       //Move FIRE HMW
       //H1
       "M256_Manag_IDB".M256F_IDB[0].tHMW.dHeadFireONReaction_ms := "DB_M256F_Scada".tHMW.dHeadFireONReaction_ms_H1;
       "M256_Manag_IDB".M256F_IDB[0].tHMW.dHeadFireOFFReaction_ms := "DB_M256F_Scada".tHMW.dHeadFireOFFReaction_ms_H1;
       "M256_Manag_IDB".M256F_IDB[0].tHMW.dHeadOilONDelay_ms := "DB_M256F_Scada".tHMW.dHeadOilONDelay_ms_H1;
       "M256_Manag_IDB".M256F_IDB[0].tHMW.dHeadOilOFFDelay_ms := "DB_M256F_Scada".tHMW.dHeadOilOFFDelay_ms_H1;
       "M256_Manag_IDB".M256F_IDB[0].tHMW.dHeadFireONDelay_cmm := "DB_M256F_Scada".tHMW.dHeadFireONDelay_cmm_H1;
       "M256_Manag_IDB".M256F_IDB[0].tHMW.dHeadFireOFFDelay_cmm := "DB_M256F_Scada".tHMW.dHeadFireOFFDelay_cmm_H1;
       "M256_Manag_IDB".M256F_IDB[0].tHMW.dHeadPressure_mN := "DB_M256F_Scada".tHMW.dHeadPressure_mN_H1;
       "M256_Manag_IDB".M256F_IDB[0].tHMW.xResetUsageCounter := "DB_M256F_Scada".tHMW.xResetUsageCounter_H1;
       "M256_Manag_IDB".M256F_IDB[0].tHMW.tManCmd.xMan_FireON := "DB_M256F_Scada".tHMW.tManCmd.xMan_FireON_H1;
       "M256_Manag_IDB".M256F_IDB[0].tHMW.tManCmd.xMan_FireOFF := "DB_M256F_Scada".tHMW.tManCmd.xMan_FireOFF_H1;
       "M256_Manag_IDB".M256F_IDB[0].tHMW.tManCmd.xMan_OilON := "DB_M256F_Scada".tHMW.tManCmd.xMan_OilON_H1;
       //H2
       "M256_Manag_IDB".M256F_IDB[1].tHMW.dHeadFireONReaction_ms := "DB_M256F_Scada".tHMW.dHeadFireONReaction_ms_H2;
       "M256_Manag_IDB".M256F_IDB[1].tHMW.dHeadFireOFFReaction_ms := "DB_M256F_Scada".tHMW.dHeadFireOFFReaction_ms_H2;
       "M256_Manag_IDB".M256F_IDB[1].tHMW.dHeadOilONDelay_ms := "DB_M256F_Scada".tHMW.dHeadOilONDelay_ms_H2;
       "M256_Manag_IDB".M256F_IDB[1].tHMW.dHeadOilOFFDelay_ms := "DB_M256F_Scada".tHMW.dHeadOilOFFDelay_ms_H2;
       "M256_Manag_IDB".M256F_IDB[1].tHMW.dHeadFireONDelay_cmm := "DB_M256F_Scada".tHMW.dHeadFireONDelay_cmm_H2;
       "M256_Manag_IDB".M256F_IDB[1].tHMW.dHeadFireOFFDelay_cmm := "DB_M256F_Scada".tHMW.dHeadFireOFFDelay_cmm_H2;
       "M256_Manag_IDB".M256F_IDB[1].tHMW.dHeadPressure_mN := "DB_M256F_Scada".tHMW.dHeadPressure_mN_H2;
       "M256_Manag_IDB".M256F_IDB[1].tHMW.xResetUsageCounter := "DB_M256F_Scada".tHMW.xResetUsageCounter_H2;
       "M256_Manag_IDB".M256F_IDB[1].tHMW.tManCmd.xMan_FireON := "DB_M256F_Scada".tHMW.tManCmd.xMan_FireON_H2;
       "M256_Manag_IDB".M256F_IDB[1].tHMW.tManCmd.xMan_FireOFF := "DB_M256F_Scada".tHMW.tManCmd.xMan_FireOFF_H2;
       "M256_Manag_IDB".M256F_IDB[1].tHMW.tManCmd.xMan_OilON := "DB_M256F_Scada".tHMW.tManCmd.xMan_OilON_H2;
       //H3
       "M256_Manag_IDB".M256F_IDB[2].tHMW.dHeadFireONReaction_ms := "DB_M256F_Scada".tHMW.dHeadFireONReaction_ms_H3;
       "M256_Manag_IDB".M256F_IDB[2].tHMW.dHeadFireOFFReaction_ms := "DB_M256F_Scada".tHMW.dHeadFireOFFReaction_ms_H3;
       "M256_Manag_IDB".M256F_IDB[2].tHMW.dHeadOilONDelay_ms := "DB_M256F_Scada".tHMW.dHeadOilONDelay_ms_H3;
       "M256_Manag_IDB".M256F_IDB[2].tHMW.dHeadOilOFFDelay_ms := "DB_M256F_Scada".tHMW.dHeadOilOFFDelay_ms_H3;
       "M256_Manag_IDB".M256F_IDB[2].tHMW.dHeadFireONDelay_cmm := "DB_M256F_Scada".tHMW.dHeadFireONDelay_cmm_H3;
       "M256_Manag_IDB".M256F_IDB[2].tHMW.dHeadFireOFFDelay_cmm := "DB_M256F_Scada".tHMW.dHeadFireOFFDelay_cmm_H3;
       "M256_Manag_IDB".M256F_IDB[2].tHMW.dHeadPressure_mN := "DB_M256F_Scada".tHMW.dHeadPressure_mN_H3;
       "M256_Manag_IDB".M256F_IDB[2].tHMW.xResetUsageCounter := "DB_M256F_Scada".tHMW.xResetUsageCounter_H3;
       "M256_Manag_IDB".M256F_IDB[2].tHMW.tManCmd.xMan_FireON := "DB_M256F_Scada".tHMW.tManCmd.xMan_FireON_H3;
       "M256_Manag_IDB".M256F_IDB[2].tHMW.tManCmd.xMan_FireOFF := "DB_M256F_Scada".tHMW.tManCmd.xMan_FireOFF_H3;
       "M256_Manag_IDB".M256F_IDB[2].tHMW.tManCmd.xMan_OilON := "DB_M256F_Scada".tHMW.tManCmd.xMan_OilON_H3;
       //H4
       "M256_Manag_IDB".M256F_IDB[3].tHMW.dHeadFireONReaction_ms := "DB_M256F_Scada".tHMW.dHeadFireONReaction_ms_H4;
       "M256_Manag_IDB".M256F_IDB[3].tHMW.dHeadFireOFFReaction_ms := "DB_M256F_Scada".tHMW.dHeadFireOFFReaction_ms_H4;
       "M256_Manag_IDB".M256F_IDB[3].tHMW.dHeadOilONDelay_ms := "DB_M256F_Scada".tHMW.dHeadOilONDelay_ms_H4;
       "M256_Manag_IDB".M256F_IDB[3].tHMW.dHeadOilOFFDelay_ms := "DB_M256F_Scada".tHMW.dHeadOilOFFDelay_ms_H4;
       "M256_Manag_IDB".M256F_IDB[3].tHMW.dHeadFireONDelay_cmm := "DB_M256F_Scada".tHMW.dHeadFireONDelay_cmm_H4;
       "M256_Manag_IDB".M256F_IDB[3].tHMW.dHeadFireOFFDelay_cmm := "DB_M256F_Scada".tHMW.dHeadFireOFFDelay_cmm_H4;
       "M256_Manag_IDB".M256F_IDB[3].tHMW.dHeadPressure_mN := "DB_M256F_Scada".tHMW.dHeadPressure_mN_H4;
       "M256_Manag_IDB".M256F_IDB[3].tHMW.xResetUsageCounter := "DB_M256F_Scada".tHMW.xResetUsageCounter_H4;
       "M256_Manag_IDB".M256F_IDB[3].tHMW.tManCmd.xMan_FireON := "DB_M256F_Scada".tHMW.tManCmd.xMan_FireON_H4;
       "M256_Manag_IDB".M256F_IDB[3].tHMW.tManCmd.xMan_FireOFF := "DB_M256F_Scada".tHMW.tManCmd.xMan_FireOFF_H4;
       "M256_Manag_IDB".M256F_IDB[3].tHMW.tManCmd.xMan_OilON := "DB_M256F_Scada".tHMW.tManCmd.xMan_OilON_H4;
       //H5
       "M256_Manag_IDB".M256F_IDB[4].tHMW.dHeadFireONReaction_ms := "DB_M256F_Scada".tHMW.dHeadFireONReaction_ms_H5;
       "M256_Manag_IDB".M256F_IDB[4].tHMW.dHeadFireOFFReaction_ms := "DB_M256F_Scada".tHMW.dHeadFireOFFReaction_ms_H5;
       "M256_Manag_IDB".M256F_IDB[4].tHMW.dHeadOilONDelay_ms := "DB_M256F_Scada".tHMW.dHeadOilONDelay_ms_H5;
       "M256_Manag_IDB".M256F_IDB[4].tHMW.dHeadOilOFFDelay_ms := "DB_M256F_Scada".tHMW.dHeadOilOFFDelay_ms_H5;
       "M256_Manag_IDB".M256F_IDB[4].tHMW.dHeadFireONDelay_cmm := "DB_M256F_Scada".tHMW.dHeadFireONDelay_cmm_H5;
       "M256_Manag_IDB".M256F_IDB[4].tHMW.dHeadFireOFFDelay_cmm := "DB_M256F_Scada".tHMW.dHeadFireOFFDelay_cmm_H5;
       "M256_Manag_IDB".M256F_IDB[4].tHMW.dHeadPressure_mN := "DB_M256F_Scada".tHMW.dHeadPressure_mN_H5;
       "M256_Manag_IDB".M256F_IDB[4].tHMW.xResetUsageCounter := "DB_M256F_Scada".tHMW.xResetUsageCounter_H5;
       "M256_Manag_IDB".M256F_IDB[4].tHMW.tManCmd.xMan_FireON := "DB_M256F_Scada".tHMW.tManCmd.xMan_FireON_H5;
       "M256_Manag_IDB".M256F_IDB[4].tHMW.tManCmd.xMan_FireOFF := "DB_M256F_Scada".tHMW.tManCmd.xMan_FireOFF_H5;
       "M256_Manag_IDB".M256F_IDB[4].tHMW.tManCmd.xMan_OilON := "DB_M256F_Scada".tHMW.tManCmd.xMan_OilON_H5;
       //H6
       "M256_Manag_IDB".M256F_IDB[5].tHMW.dHeadFireONReaction_ms := "DB_M256F_Scada".tHMW.dHeadFireONReaction_ms_H6;
       "M256_Manag_IDB".M256F_IDB[5].tHMW.dHeadFireOFFReaction_ms := "DB_M256F_Scada".tHMW.dHeadFireOFFReaction_ms_H6;
       "M256_Manag_IDB".M256F_IDB[5].tHMW.dHeadOilONDelay_ms := "DB_M256F_Scada".tHMW.dHeadOilONDelay_ms_H6;
       "M256_Manag_IDB".M256F_IDB[5].tHMW.dHeadOilOFFDelay_ms := "DB_M256F_Scada".tHMW.dHeadOilOFFDelay_ms_H6;
       "M256_Manag_IDB".M256F_IDB[5].tHMW.dHeadFireONDelay_cmm := "DB_M256F_Scada".tHMW.dHeadFireONDelay_cmm_H6;
       "M256_Manag_IDB".M256F_IDB[5].tHMW.dHeadFireOFFDelay_cmm := "DB_M256F_Scada".tHMW.dHeadFireOFFDelay_cmm_H6;
       "M256_Manag_IDB".M256F_IDB[5].tHMW.dHeadPressure_mN := "DB_M256F_Scada".tHMW.dHeadPressure_mN_H6;
       "M256_Manag_IDB".M256F_IDB[5].tHMW.xResetUsageCounter := "DB_M256F_Scada".tHMW.xResetUsageCounter_H6;
       "M256_Manag_IDB".M256F_IDB[5].tHMW.tManCmd.xMan_FireON := "DB_M256F_Scada".tHMW.tManCmd.xMan_FireON_H6;
       "M256_Manag_IDB".M256F_IDB[5].tHMW.tManCmd.xMan_FireOFF := "DB_M256F_Scada".tHMW.tManCmd.xMan_FireOFF_H6;
       "M256_Manag_IDB".M256F_IDB[5].tHMW.tManCmd.xMan_OilON := "DB_M256F_Scada".tHMW.tManCmd.xMan_OilON_H6;
       //H7
       "M256_Manag_IDB".M256F_IDB[6].tHMW.dHeadFireONReaction_ms := "DB_M256F_Scada".tHMW.dHeadFireONReaction_ms_H7;
       "M256_Manag_IDB".M256F_IDB[6].tHMW.dHeadFireOFFReaction_ms := "DB_M256F_Scada".tHMW.dHeadFireOFFReaction_ms_H7;
       "M256_Manag_IDB".M256F_IDB[6].tHMW.dHeadOilONDelay_ms := "DB_M256F_Scada".tHMW.dHeadOilONDelay_ms_H7;
       "M256_Manag_IDB".M256F_IDB[6].tHMW.dHeadOilOFFDelay_ms := "DB_M256F_Scada".tHMW.dHeadOilOFFDelay_ms_H7;
       "M256_Manag_IDB".M256F_IDB[6].tHMW.dHeadFireONDelay_cmm := "DB_M256F_Scada".tHMW.dHeadFireONDelay_cmm_H7;
       "M256_Manag_IDB".M256F_IDB[6].tHMW.dHeadFireOFFDelay_cmm := "DB_M256F_Scada".tHMW.dHeadFireOFFDelay_cmm_H7;
       "M256_Manag_IDB".M256F_IDB[6].tHMW.dHeadPressure_mN := "DB_M256F_Scada".tHMW.dHeadPressure_mN_H7;
       "M256_Manag_IDB".M256F_IDB[6].tHMW.xResetUsageCounter := "DB_M256F_Scada".tHMW.xResetUsageCounter_H7;
       "M256_Manag_IDB".M256F_IDB[6].tHMW.tManCmd.xMan_FireON := "DB_M256F_Scada".tHMW.tManCmd.xMan_FireON_H7;
       "M256_Manag_IDB".M256F_IDB[6].tHMW.tManCmd.xMan_FireOFF := "DB_M256F_Scada".tHMW.tManCmd.xMan_FireOFF_H7;
       "M256_Manag_IDB".M256F_IDB[6].tHMW.tManCmd.xMan_OilON := "DB_M256F_Scada".tHMW.tManCmd.xMan_OilON_H7;
       //H8
       "M256_Manag_IDB".M256F_IDB[7].tHMW.dHeadFireONReaction_ms := "DB_M256F_Scada".tHMW.dHeadFireONReaction_ms_H8;
       "M256_Manag_IDB".M256F_IDB[7].tHMW.dHeadFireOFFReaction_ms := "DB_M256F_Scada".tHMW.dHeadFireOFFReaction_ms_H8;
       "M256_Manag_IDB".M256F_IDB[7].tHMW.dHeadOilONDelay_ms := "DB_M256F_Scada".tHMW.dHeadOilONDelay_ms_H8;
       "M256_Manag_IDB".M256F_IDB[7].tHMW.dHeadOilOFFDelay_ms := "DB_M256F_Scada".tHMW.dHeadOilOFFDelay_ms_H8;
       "M256_Manag_IDB".M256F_IDB[7].tHMW.dHeadFireONDelay_cmm := "DB_M256F_Scada".tHMW.dHeadFireONDelay_cmm_H8;
       "M256_Manag_IDB".M256F_IDB[7].tHMW.dHeadFireOFFDelay_cmm := "DB_M256F_Scada".tHMW.dHeadFireOFFDelay_cmm_H8;
       "M256_Manag_IDB".M256F_IDB[7].tHMW.dHeadPressure_mN := "DB_M256F_Scada".tHMW.dHeadPressure_mN_H8;
       "M256_Manag_IDB".M256F_IDB[7].tHMW.xResetUsageCounter := "DB_M256F_Scada".tHMW.xResetUsageCounter_H8;
       "M256_Manag_IDB".M256F_IDB[7].tHMW.tManCmd.xMan_FireON := "DB_M256F_Scada".tHMW.tManCmd.xMan_FireON_H8;
       "M256_Manag_IDB".M256F_IDB[7].tHMW.tManCmd.xMan_FireOFF := "DB_M256F_Scada".tHMW.tManCmd.xMan_FireOFF_H8;
       "M256_Manag_IDB".M256F_IDB[7].tHMW.tManCmd.xMan_OilON := "DB_M256F_Scada".tHMW.tManCmd.xMan_OilON_H8;

       //Move FIRE ALM
       "DB_M256F_Scada".tAlm.tF:="M256_Manag_IDB".M256F_IDB[0].tALM.tF;

       "DB_M256F_Scada".tAlm.tW := "M256_Manag_IDB".M256F_IDB[0].tALM.tW;

       //H1
       "DB_M256F_Scada".tAlm.tS.tS0.x0 := "M256_Manag_IDB".M256F_IDB[0].tALM.tS.x0;
       "DB_M256F_Scada".tAlm.tS.tS0.x1 := "M256_Manag_IDB".M256F_IDB[0].tALM.tS.x1;
       "DB_M256F_Scada".tAlm.tS.tS0.x2 := "M256_Manag_IDB".M256F_IDB[0].tALM.tS.x2;
       "DB_M256F_Scada".tAlm.tS.tS0.x3 := "M256_Manag_IDB".M256F_IDB[0].tALM.tS.x3;
       "DB_M256F_Scada".tAlm.tS.tS0.x4 := "M256_Manag_IDB".M256F_IDB[0].tALM.tS.x4;
       "DB_M256F_Scada".tAlm.tS.tS0.x5 := "M256_Manag_IDB".M256F_IDB[0].tALM.tS.x5;
       "DB_M256F_Scada".tAlm.tS.tS0.x6 := "M256_Manag_IDB".M256F_IDB[0].tALM.tS.x6;
       "DB_M256F_Scada".tAlm.tS.tS0.x7 := "M256_Manag_IDB".M256F_IDB[0].tALM.tS.x7;
       "DB_M256F_Scada".tAlm.tS.tS0.x8 := "M256_Manag_IDB".M256F_IDB[0].tALM.tS.x8;
       //H2
       "DB_M256F_Scada".tAlm.tS.tS0.x9 := "M256_Manag_IDB".M256F_IDB[1].tALM.tS.x0;
       "DB_M256F_Scada".tAlm.tS.tS0.x10 := "M256_Manag_IDB".M256F_IDB[1].tALM.tS.x1;
       "DB_M256F_Scada".tAlm.tS.tS0.x11 := "M256_Manag_IDB".M256F_IDB[1].tALM.tS.x2;
       "DB_M256F_Scada".tAlm.tS.tS0.x12 := "M256_Manag_IDB".M256F_IDB[1].tALM.tS.x3;
       "DB_M256F_Scada".tAlm.tS.tS0.x13 := "M256_Manag_IDB".M256F_IDB[1].tALM.tS.x4;
       "DB_M256F_Scada".tAlm.tS.tS0.x14 := "M256_Manag_IDB".M256F_IDB[1].tALM.tS.x5;
       "DB_M256F_Scada".tAlm.tS.tS0.x15 := "M256_Manag_IDB".M256F_IDB[1].tALM.tS.x6;
       "DB_M256F_Scada".tAlm.tS.tS0.x16 := "M256_Manag_IDB".M256F_IDB[1].tALM.tS.x7;
       "DB_M256F_Scada".tAlm.tS.tS0.x17 := "M256_Manag_IDB".M256F_IDB[1].tALM.tS.x8;
       //H3
       "DB_M256F_Scada".tAlm.tS.tS0.x18 := "M256_Manag_IDB".M256F_IDB[2].tALM.tS.x0;
       "DB_M256F_Scada".tAlm.tS.tS0.x19 := "M256_Manag_IDB".M256F_IDB[2].tALM.tS.x1;
       "DB_M256F_Scada".tAlm.tS.tS0.x20 := "M256_Manag_IDB".M256F_IDB[2].tALM.tS.x2;
       "DB_M256F_Scada".tAlm.tS.tS0.x21 := "M256_Manag_IDB".M256F_IDB[2].tALM.tS.x3;
       "DB_M256F_Scada".tAlm.tS.tS0.x22 := "M256_Manag_IDB".M256F_IDB[2].tALM.tS.x4;
       "DB_M256F_Scada".tAlm.tS.tS0.x23 := "M256_Manag_IDB".M256F_IDB[2].tALM.tS.x5;
       "DB_M256F_Scada".tAlm.tS.tS0.x24 := "M256_Manag_IDB".M256F_IDB[2].tALM.tS.x6;
       "DB_M256F_Scada".tAlm.tS.tS0.x25 := "M256_Manag_IDB".M256F_IDB[2].tALM.tS.x7;
       "DB_M256F_Scada".tAlm.tS.tS0.x26 := "M256_Manag_IDB".M256F_IDB[2].tALM.tS.x8;
       //H4
       "DB_M256F_Scada".tAlm.tS.tS1.x0 := "M256_Manag_IDB".M256F_IDB[3].tALM.tS.x0;
       "DB_M256F_Scada".tAlm.tS.tS1.x1 := "M256_Manag_IDB".M256F_IDB[3].tALM.tS.x1;
       "DB_M256F_Scada".tAlm.tS.tS1.x2 := "M256_Manag_IDB".M256F_IDB[3].tALM.tS.x2;
       "DB_M256F_Scada".tAlm.tS.tS1.x3 := "M256_Manag_IDB".M256F_IDB[3].tALM.tS.x3;
       "DB_M256F_Scada".tAlm.tS.tS1.x4 := "M256_Manag_IDB".M256F_IDB[3].tALM.tS.x4;
       "DB_M256F_Scada".tAlm.tS.tS1.x5 := "M256_Manag_IDB".M256F_IDB[3].tALM.tS.x5;
       "DB_M256F_Scada".tAlm.tS.tS1.x6 := "M256_Manag_IDB".M256F_IDB[3].tALM.tS.x6;
       "DB_M256F_Scada".tAlm.tS.tS1.x7 := "M256_Manag_IDB".M256F_IDB[3].tALM.tS.x7;
       "DB_M256F_Scada".tAlm.tS.tS1.x8 := "M256_Manag_IDB".M256F_IDB[3].tALM.tS.x8;
       //H5
       "DB_M256F_Scada".tAlm.tS.tS1.x9 := "M256_Manag_IDB".M256F_IDB[4].tALM.tS.x0;
       "DB_M256F_Scada".tAlm.tS.tS1.x10 := "M256_Manag_IDB".M256F_IDB[4].tALM.tS.x1;
       "DB_M256F_Scada".tAlm.tS.tS1.x11 := "M256_Manag_IDB".M256F_IDB[4].tALM.tS.x2;
       "DB_M256F_Scada".tAlm.tS.tS1.x12 := "M256_Manag_IDB".M256F_IDB[4].tALM.tS.x3;
       "DB_M256F_Scada".tAlm.tS.tS1.x13 := "M256_Manag_IDB".M256F_IDB[4].tALM.tS.x4;
       "DB_M256F_Scada".tAlm.tS.tS1.x14 := "M256_Manag_IDB".M256F_IDB[4].tALM.tS.x5;
       "DB_M256F_Scada".tAlm.tS.tS1.x15 := "M256_Manag_IDB".M256F_IDB[4].tALM.tS.x6;
       "DB_M256F_Scada".tAlm.tS.tS1.x16 := "M256_Manag_IDB".M256F_IDB[4].tALM.tS.x7;
       "DB_M256F_Scada".tAlm.tS.tS1.x17 := "M256_Manag_IDB".M256F_IDB[4].tALM.tS.x8;
       //H6
       "DB_M256F_Scada".tAlm.tS.tS1.x18 := "M256_Manag_IDB".M256F_IDB[5].tALM.tS.x0;
       "DB_M256F_Scada".tAlm.tS.tS1.x19 := "M256_Manag_IDB".M256F_IDB[5].tALM.tS.x1;
       "DB_M256F_Scada".tAlm.tS.tS1.x20 := "M256_Manag_IDB".M256F_IDB[5].tALM.tS.x2;
       "DB_M256F_Scada".tAlm.tS.tS1.x21 := "M256_Manag_IDB".M256F_IDB[5].tALM.tS.x3;
       "DB_M256F_Scada".tAlm.tS.tS1.x22 := "M256_Manag_IDB".M256F_IDB[5].tALM.tS.x4;
       "DB_M256F_Scada".tAlm.tS.tS1.x23 := "M256_Manag_IDB".M256F_IDB[5].tALM.tS.x5;
       "DB_M256F_Scada".tAlm.tS.tS1.x24 := "M256_Manag_IDB".M256F_IDB[5].tALM.tS.x6;
       "DB_M256F_Scada".tAlm.tS.tS1.x25 := "M256_Manag_IDB".M256F_IDB[5].tALM.tS.x7;
       "DB_M256F_Scada".tAlm.tS.tS1.x26 := "M256_Manag_IDB".M256F_IDB[5].tALM.tS.x8;
       //H7
       "DB_M256F_Scada".tAlm.tS.tS2.x0 := "M256_Manag_IDB".M256F_IDB[6].tALM.tS.x0;
       "DB_M256F_Scada".tAlm.tS.tS2.x1 := "M256_Manag_IDB".M256F_IDB[6].tALM.tS.x1;
       "DB_M256F_Scada".tAlm.tS.tS2.x2 := "M256_Manag_IDB".M256F_IDB[6].tALM.tS.x2;
       "DB_M256F_Scada".tAlm.tS.tS2.x3 := "M256_Manag_IDB".M256F_IDB[6].tALM.tS.x3;
       "DB_M256F_Scada".tAlm.tS.tS2.x4 := "M256_Manag_IDB".M256F_IDB[6].tALM.tS.x4;
       "DB_M256F_Scada".tAlm.tS.tS2.x5 := "M256_Manag_IDB".M256F_IDB[6].tALM.tS.x5;
       "DB_M256F_Scada".tAlm.tS.tS2.x6 := "M256_Manag_IDB".M256F_IDB[6].tALM.tS.x6;
       "DB_M256F_Scada".tAlm.tS.tS2.x7 := "M256_Manag_IDB".M256F_IDB[6].tALM.tS.x7;
       "DB_M256F_Scada".tAlm.tS.tS2.x8 := "M256_Manag_IDB".M256F_IDB[6].tALM.tS.x8;
       //H8
       "DB_M256F_Scada".tAlm.tS.tS2.x9 := "M256_Manag_IDB".M256F_IDB[7].tALM.tS.x0;
       "DB_M256F_Scada".tAlm.tS.tS2.x10 := "M256_Manag_IDB".M256F_IDB[7].tALM.tS.x1;
       "DB_M256F_Scada".tAlm.tS.tS2.x11 := "M256_Manag_IDB".M256F_IDB[7].tALM.tS.x2;
       "DB_M256F_Scada".tAlm.tS.tS2.x12 := "M256_Manag_IDB".M256F_IDB[7].tALM.tS.x3;
       "DB_M256F_Scada".tAlm.tS.tS2.x13 := "M256_Manag_IDB".M256F_IDB[7].tALM.tS.x4;
       "DB_M256F_Scada".tAlm.tS.tS2.x14 := "M256_Manag_IDB".M256F_IDB[7].tALM.tS.x5;
       "DB_M256F_Scada".tAlm.tS.tS2.x15 := "M256_Manag_IDB".M256F_IDB[7].tALM.tS.x6;
       "DB_M256F_Scada".tAlm.tS.tS2.x16 := "M256_Manag_IDB".M256F_IDB[7].tALM.tS.x7;
       "DB_M256F_Scada".tAlm.tS.tS2.x17 := "M256_Manag_IDB".M256F_IDB[7].tALM.tS.x8;



       //Move ARMING HMR
       //H1
       "DB_M256A_Scada".tHMR.dHeadStatus_H1 := "M256_Manag_IDB".M256A_IDB[0].tHMR.dHeadStatus;
       "DB_M256A_Scada".tHMR.tManCmd.xMan_DescentFdbk_H1:="M256_Manag_IDB".M256A_IDB[0].tHMR.tManCmd.xMan_DescentFdbk;
       "DB_M256A_Scada".tHMR.tManCmd.xMan_RiseFdbk_H1 := "M256_Manag_IDB".M256A_IDB[0].tHMR.tManCmd.xMan_RiseFdbk;
       //H2
       "DB_M256A_Scada".tHMR.dHeadStatus_H2 := "M256_Manag_IDB".M256A_IDB[1].tHMR.dHeadStatus;
       "DB_M256A_Scada".tHMR.tManCmd.xMan_DescentFdbk_H2 := "M256_Manag_IDB".M256A_IDB[1].tHMR.tManCmd.xMan_DescentFdbk;
       "DB_M256A_Scada".tHMR.tManCmd.xMan_RiseFdbk_H2 := "M256_Manag_IDB".M256A_IDB[1].tHMR.tManCmd.xMan_RiseFdbk;
       //H3
       "DB_M256A_Scada".tHMR.dHeadStatus_H3 := "M256_Manag_IDB".M256A_IDB[2].tHMR.dHeadStatus;
       "DB_M256A_Scada".tHMR.tManCmd.xMan_DescentFdbk_H3 := "M256_Manag_IDB".M256A_IDB[2].tHMR.tManCmd.xMan_DescentFdbk;
       "DB_M256A_Scada".tHMR.tManCmd.xMan_RiseFdbk_H3 := "M256_Manag_IDB".M256A_IDB[2].tHMR.tManCmd.xMan_RiseFdbk;
       //H4
       "DB_M256A_Scada".tHMR.dHeadStatus_H4 := "M256_Manag_IDB".M256A_IDB[3].tHMR.dHeadStatus;
       "DB_M256A_Scada".tHMR.tManCmd.xMan_DescentFdbk_H4 := "M256_Manag_IDB".M256A_IDB[3].tHMR.tManCmd.xMan_DescentFdbk;
       "DB_M256A_Scada".tHMR.tManCmd.xMan_RiseFdbk_H4 := "M256_Manag_IDB".M256A_IDB[3].tHMR.tManCmd.xMan_RiseFdbk;
       //H5
       "DB_M256A_Scada".tHMR.dHeadStatus_H5 := "M256_Manag_IDB".M256A_IDB[4].tHMR.dHeadStatus;
       "DB_M256A_Scada".tHMR.tManCmd.xMan_DescentFdbk_H5 := "M256_Manag_IDB".M256A_IDB[4].tHMR.tManCmd.xMan_DescentFdbk;
       "DB_M256A_Scada".tHMR.tManCmd.xMan_RiseFdbk_H5 := "M256_Manag_IDB".M256A_IDB[4].tHMR.tManCmd.xMan_RiseFdbk;
       //H6
       "DB_M256A_Scada".tHMR.dHeadStatus_H6 := "M256_Manag_IDB".M256A_IDB[5].tHMR.dHeadStatus;
       "DB_M256A_Scada".tHMR.tManCmd.xMan_DescentFdbk_H6 := "M256_Manag_IDB".M256A_IDB[5].tHMR.tManCmd.xMan_DescentFdbk;
       "DB_M256A_Scada".tHMR.tManCmd.xMan_RiseFdbk_H6 := "M256_Manag_IDB".M256A_IDB[5].tHMR.tManCmd.xMan_RiseFdbk;
       //H7
       "DB_M256A_Scada".tHMR.dHeadStatus_H7 := "M256_Manag_IDB".M256A_IDB[6].tHMR.dHeadStatus;
       "DB_M256A_Scada".tHMR.tManCmd.xMan_DescentFdbk_H7 := "M256_Manag_IDB".M256A_IDB[6].tHMR.tManCmd.xMan_DescentFdbk;
       "DB_M256A_Scada".tHMR.tManCmd.xMan_RiseFdbk_H7 := "M256_Manag_IDB".M256A_IDB[6].tHMR.tManCmd.xMan_RiseFdbk;
       //H8
       "DB_M256A_Scada".tHMR.dHeadStatus_H8 := "M256_Manag_IDB".M256A_IDB[7].tHMR.dHeadStatus;
       "DB_M256A_Scada".tHMR.tManCmd.xMan_DescentFdbk_H8 := "M256_Manag_IDB".M256A_IDB[7].tHMR.tManCmd.xMan_DescentFdbk;
       "DB_M256A_Scada".tHMR.tManCmd.xMan_RiseFdbk_H8 := "M256_Manag_IDB".M256A_IDB[7].tHMR.tManCmd.xMan_RiseFdbk;

       //Move ARMING HMW
       //H1
       "M256_Manag_IDB".M256A_IDB[0].tHMW.dDescentReactTime_ms:="DB_M256A_Scada".tHMW.dDescentReactTime_ms_H1;
       "M256_Manag_IDB".M256A_IDB[0].tHMW.dRaiseReactTime_ms := "DB_M256A_Scada".tHMW.dRaiseReactTime_ms_H1;
       "M256_Manag_IDB".M256A_IDB[0].tHMW.tManCmd.xManDescent := "DB_M256A_Scada".tHMW.tManCmd.xManDescent_H1;
       "M256_Manag_IDB".M256A_IDB[0].tHMW.tManCmd.xManRise := "DB_M256A_Scada".tHMW.tManCmd.xManRise_H1;
       //H2
       "M256_Manag_IDB".M256A_IDB[1].tHMW.dDescentReactTime_ms := "DB_M256A_Scada".tHMW.dDescentReactTime_ms_H2;
       "M256_Manag_IDB".M256A_IDB[1].tHMW.dRaiseReactTime_ms := "DB_M256A_Scada".tHMW.dRaiseReactTime_ms_H2;
       "M256_Manag_IDB".M256A_IDB[1].tHMW.tManCmd.xManDescent := "DB_M256A_Scada".tHMW.tManCmd.xManDescent_H2;
       "M256_Manag_IDB".M256A_IDB[1].tHMW.tManCmd.xManRise := "DB_M256A_Scada".tHMW.tManCmd.xManRise_H2;
       //H3
       "M256_Manag_IDB".M256A_IDB[2].tHMW.dDescentReactTime_ms := "DB_M256A_Scada".tHMW.dDescentReactTime_ms_H3;
       "M256_Manag_IDB".M256A_IDB[2].tHMW.dRaiseReactTime_ms := "DB_M256A_Scada".tHMW.dRaiseReactTime_ms_H3;
       "M256_Manag_IDB".M256A_IDB[2].tHMW.tManCmd.xManDescent := "DB_M256A_Scada".tHMW.tManCmd.xManDescent_H3;
       "M256_Manag_IDB".M256A_IDB[2].tHMW.tManCmd.xManRise := "DB_M256A_Scada".tHMW.tManCmd.xManRise_H3;
       //H4
       "M256_Manag_IDB".M256A_IDB[3].tHMW.dDescentReactTime_ms := "DB_M256A_Scada".tHMW.dDescentReactTime_ms_H4;
       "M256_Manag_IDB".M256A_IDB[3].tHMW.dRaiseReactTime_ms := "DB_M256A_Scada".tHMW.dRaiseReactTime_ms_H4;
       "M256_Manag_IDB".M256A_IDB[3].tHMW.tManCmd.xManDescent := "DB_M256A_Scada".tHMW.tManCmd.xManDescent_H4;
       "M256_Manag_IDB".M256A_IDB[3].tHMW.tManCmd.xManRise := "DB_M256A_Scada".tHMW.tManCmd.xManRise_H4;
       //H5
       "M256_Manag_IDB".M256A_IDB[4].tHMW.dDescentReactTime_ms := "DB_M256A_Scada".tHMW.dDescentReactTime_ms_H5;
       "M256_Manag_IDB".M256A_IDB[4].tHMW.dRaiseReactTime_ms := "DB_M256A_Scada".tHMW.dRaiseReactTime_ms_H5;
       "M256_Manag_IDB".M256A_IDB[4].tHMW.tManCmd.xManDescent := "DB_M256A_Scada".tHMW.tManCmd.xManDescent_H5;
       "M256_Manag_IDB".M256A_IDB[4].tHMW.tManCmd.xManRise := "DB_M256A_Scada".tHMW.tManCmd.xManRise_H5;
       //H6
       "M256_Manag_IDB".M256A_IDB[5].tHMW.dDescentReactTime_ms := "DB_M256A_Scada".tHMW.dDescentReactTime_ms_H6;
       "M256_Manag_IDB".M256A_IDB[5].tHMW.dRaiseReactTime_ms := "DB_M256A_Scada".tHMW.dRaiseReactTime_ms_H6;
       "M256_Manag_IDB".M256A_IDB[5].tHMW.tManCmd.xManDescent := "DB_M256A_Scada".tHMW.tManCmd.xManDescent_H6;
       "M256_Manag_IDB".M256A_IDB[5].tHMW.tManCmd.xManRise := "DB_M256A_Scada".tHMW.tManCmd.xManRise_H6;
       //H7
       "M256_Manag_IDB".M256A_IDB[6].tHMW.dDescentReactTime_ms := "DB_M256A_Scada".tHMW.dDescentReactTime_ms_H7;
       "M256_Manag_IDB".M256A_IDB[6].tHMW.dRaiseReactTime_ms := "DB_M256A_Scada".tHMW.dRaiseReactTime_ms_H7;
       "M256_Manag_IDB".M256A_IDB[6].tHMW.tManCmd.xManDescent := "DB_M256A_Scada".tHMW.tManCmd.xManDescent_H7;
       "M256_Manag_IDB".M256A_IDB[6].tHMW.tManCmd.xManRise := "DB_M256A_Scada".tHMW.tManCmd.xManRise_H7;
       //H8
       "M256_Manag_IDB".M256A_IDB[7].tHMW.dDescentReactTime_ms := "DB_M256A_Scada".tHMW.dDescentReactTime_ms_H8;
       "M256_Manag_IDB".M256A_IDB[7].tHMW.dRaiseReactTime_ms := "DB_M256A_Scada".tHMW.dRaiseReactTime_ms_H8;
       "M256_Manag_IDB".M256A_IDB[7].tHMW.tManCmd.xManDescent := "DB_M256A_Scada".tHMW.tManCmd.xManDescent_H8;
       "M256_Manag_IDB".M256A_IDB[7].tHMW.tManCmd.xManRise := "DB_M256A_Scada".tHMW.tManCmd.xManRise_H8;


       //Move ARMING ALM

       "DB_M256A_Scada".tAlm.tF := "M256_Manag_IDB".M256A_IDB[0].tALM.tF;

       "DB_M256A_Scada".tAlm.tW := "M256_Manag_IDB".M256A_IDB[0].tALM.tW;

               //H1
       "DB_M256A_Scada".tAlm.tS.tS0.x0 := "M256_Manag_IDB".M256A_IDB[0].tALM.tS.xNotWorkPos;
       "DB_M256A_Scada".tAlm.tS.tS0.x1 := "M256_Manag_IDB".M256A_IDB[0].tALM.tS.x1;
       "DB_M256A_Scada".tAlm.tS.tS0.x2 := "M256_Manag_IDB".M256A_IDB[0].tALM.tS.x2;
       "DB_M256A_Scada".tAlm.tS.tS0.x3 := "M256_Manag_IDB".M256A_IDB[0].tALM.tS.x3;
       "DB_M256A_Scada".tAlm.tS.tS0.x4 := "M256_Manag_IDB".M256A_IDB[0].tALM.tS.x4;
       "DB_M256A_Scada".tAlm.tS.tS0.x5 := "M256_Manag_IDB".M256A_IDB[0].tALM.tS.x5;
       "DB_M256A_Scada".tAlm.tS.tS0.x6 := "M256_Manag_IDB".M256A_IDB[0].tALM.tS.x6;
       "DB_M256A_Scada".tAlm.tS.tS0.x7 := "M256_Manag_IDB".M256A_IDB[0].tALM.tS.x7;
       "DB_M256A_Scada".tAlm.tS.tS0.x8 := "M256_Manag_IDB".M256A_IDB[0].tALM.tS.x8;
               //H2
       "DB_M256A_Scada".tAlm.tS.tS0.x9 := "M256_Manag_IDB".M256A_IDB[1].tALM.tS.xNotWorkPos;
       "DB_M256A_Scada".tAlm.tS.tS0.x10 := "M256_Manag_IDB".M256A_IDB[1].tALM.tS.x1;
       "DB_M256A_Scada".tAlm.tS.tS0.x11 := "M256_Manag_IDB".M256A_IDB[1].tALM.tS.x2;
       "DB_M256A_Scada".tAlm.tS.tS0.x12 := "M256_Manag_IDB".M256A_IDB[1].tALM.tS.x3;
       "DB_M256A_Scada".tAlm.tS.tS0.x13 := "M256_Manag_IDB".M256A_IDB[1].tALM.tS.x4;
       "DB_M256A_Scada".tAlm.tS.tS0.x14 := "M256_Manag_IDB".M256A_IDB[1].tALM.tS.x5;
       "DB_M256A_Scada".tAlm.tS.tS0.x15 := "M256_Manag_IDB".M256A_IDB[1].tALM.tS.x6;
       "DB_M256A_Scada".tAlm.tS.tS0.x16 := "M256_Manag_IDB".M256A_IDB[1].tALM.tS.x7;
       "DB_M256A_Scada".tAlm.tS.tS0.x17 := "M256_Manag_IDB".M256A_IDB[1].tALM.tS.x8;
               //H3
       "DB_M256A_Scada".tAlm.tS.tS0.x18 := "M256_Manag_IDB".M256A_IDB[2].tALM.tS.xNotWorkPos;
       "DB_M256A_Scada".tAlm.tS.tS0.x19 := "M256_Manag_IDB".M256A_IDB[2].tALM.tS.x1;
       "DB_M256A_Scada".tAlm.tS.tS0.x20 := "M256_Manag_IDB".M256A_IDB[2].tALM.tS.x2;
       "DB_M256A_Scada".tAlm.tS.tS0.x21 := "M256_Manag_IDB".M256A_IDB[2].tALM.tS.x3;
       "DB_M256A_Scada".tAlm.tS.tS0.x22 := "M256_Manag_IDB".M256A_IDB[2].tALM.tS.x4;
       "DB_M256A_Scada".tAlm.tS.tS0.x23 := "M256_Manag_IDB".M256A_IDB[2].tALM.tS.x5;
       "DB_M256A_Scada".tAlm.tS.tS0.x24 := "M256_Manag_IDB".M256A_IDB[2].tALM.tS.x6;
       "DB_M256A_Scada".tAlm.tS.tS0.x25 := "M256_Manag_IDB".M256A_IDB[2].tALM.tS.x7;
       "DB_M256A_Scada".tAlm.tS.tS0.x26 := "M256_Manag_IDB".M256A_IDB[2].tALM.tS.x8;
               //H4
       "DB_M256A_Scada".tAlm.tS.tS1.x0 := "M256_Manag_IDB".M256A_IDB[3].tALM.tS.xNotWorkPos;
       "DB_M256A_Scada".tAlm.tS.tS1.x1 := "M256_Manag_IDB".M256A_IDB[3].tALM.tS.x1;
       "DB_M256A_Scada".tAlm.tS.tS1.x2 := "M256_Manag_IDB".M256A_IDB[3].tALM.tS.x2;
       "DB_M256A_Scada".tAlm.tS.tS1.x3 := "M256_Manag_IDB".M256A_IDB[3].tALM.tS.x3;
       "DB_M256A_Scada".tAlm.tS.tS1.x4 := "M256_Manag_IDB".M256A_IDB[3].tALM.tS.x4;
       "DB_M256A_Scada".tAlm.tS.tS1.x5 := "M256_Manag_IDB".M256A_IDB[3].tALM.tS.x5;
       "DB_M256A_Scada".tAlm.tS.tS1.x6 := "M256_Manag_IDB".M256A_IDB[3].tALM.tS.x6;
       "DB_M256A_Scada".tAlm.tS.tS1.x7 := "M256_Manag_IDB".M256A_IDB[3].tALM.tS.x7;
       "DB_M256A_Scada".tAlm.tS.tS1.x8 := "M256_Manag_IDB".M256A_IDB[3].tALM.tS.x8;
               //H5
       "DB_M256A_Scada".tAlm.tS.tS1.x9 := "M256_Manag_IDB".M256A_IDB[4].tALM.tS.xNotWorkPos;
       "DB_M256A_Scada".tAlm.tS.tS1.x10 := "M256_Manag_IDB".M256A_IDB[4].tALM.tS.x1;
       "DB_M256A_Scada".tAlm.tS.tS1.x11 := "M256_Manag_IDB".M256A_IDB[4].tALM.tS.x2;
       "DB_M256A_Scada".tAlm.tS.tS1.x12 := "M256_Manag_IDB".M256A_IDB[4].tALM.tS.x3;
       "DB_M256A_Scada".tAlm.tS.tS1.x13 := "M256_Manag_IDB".M256A_IDB[4].tALM.tS.x4;
       "DB_M256A_Scada".tAlm.tS.tS1.x14 := "M256_Manag_IDB".M256A_IDB[4].tALM.tS.x5;
       "DB_M256A_Scada".tAlm.tS.tS1.x15 := "M256_Manag_IDB".M256A_IDB[4].tALM.tS.x6;
       "DB_M256A_Scada".tAlm.tS.tS1.x16 := "M256_Manag_IDB".M256A_IDB[4].tALM.tS.x7;
       "DB_M256A_Scada".tAlm.tS.tS1.x17 := "M256_Manag_IDB".M256A_IDB[4].tALM.tS.x8;
               //H6
       "DB_M256A_Scada".tAlm.tS.tS1.x18 := "M256_Manag_IDB".M256A_IDB[5].tALM.tS.xNotWorkPos;
       "DB_M256A_Scada".tAlm.tS.tS1.x19 := "M256_Manag_IDB".M256A_IDB[5].tALM.tS.x1;
       "DB_M256A_Scada".tAlm.tS.tS1.x20 := "M256_Manag_IDB".M256A_IDB[5].tALM.tS.x2;
       "DB_M256A_Scada".tAlm.tS.tS1.x21 := "M256_Manag_IDB".M256A_IDB[5].tALM.tS.x3;
       "DB_M256A_Scada".tAlm.tS.tS1.x22 := "M256_Manag_IDB".M256A_IDB[5].tALM.tS.x4;
       "DB_M256A_Scada".tAlm.tS.tS1.x23 := "M256_Manag_IDB".M256A_IDB[5].tALM.tS.x5;
       "DB_M256A_Scada".tAlm.tS.tS1.x24 := "M256_Manag_IDB".M256A_IDB[5].tALM.tS.x6;
       "DB_M256A_Scada".tAlm.tS.tS1.x25 := "M256_Manag_IDB".M256A_IDB[5].tALM.tS.x7;
       "DB_M256A_Scada".tAlm.tS.tS1.x26 := "M256_Manag_IDB".M256A_IDB[5].tALM.tS.x8;
               //H7
       "DB_M256A_Scada".tAlm.tS.tS2.x0 := "M256_Manag_IDB".M256A_IDB[6].tALM.tS.xNotWorkPos;
       "DB_M256A_Scada".tAlm.tS.tS2.x1 := "M256_Manag_IDB".M256A_IDB[6].tALM.tS.x1;
       "DB_M256A_Scada".tAlm.tS.tS2.x2 := "M256_Manag_IDB".M256A_IDB[6].tALM.tS.x2;
       "DB_M256A_Scada".tAlm.tS.tS2.x3 := "M256_Manag_IDB".M256A_IDB[6].tALM.tS.x3;
       "DB_M256A_Scada".tAlm.tS.tS2.x4 := "M256_Manag_IDB".M256A_IDB[6].tALM.tS.x4;
       "DB_M256A_Scada".tAlm.tS.tS2.x5 := "M256_Manag_IDB".M256A_IDB[6].tALM.tS.x5;
       "DB_M256A_Scada".tAlm.tS.tS2.x6 := "M256_Manag_IDB".M256A_IDB[6].tALM.tS.x6;
       "DB_M256A_Scada".tAlm.tS.tS2.x7 := "M256_Manag_IDB".M256A_IDB[6].tALM.tS.x7;
       "DB_M256A_Scada".tAlm.tS.tS2.x8 := "M256_Manag_IDB".M256A_IDB[6].tALM.tS.x8;
               //H8
       "DB_M256A_Scada".tAlm.tS.tS2.x9 := "M256_Manag_IDB".M256A_IDB[7].tALM.tS.xNotWorkPos;
       "DB_M256A_Scada".tAlm.tS.tS2.x10 := "M256_Manag_IDB".M256A_IDB[7].tALM.tS.x1;
       "DB_M256A_Scada".tAlm.tS.tS2.x11 := "M256_Manag_IDB".M256A_IDB[7].tALM.tS.x2;
       "DB_M256A_Scada".tAlm.tS.tS2.x12 := "M256_Manag_IDB".M256A_IDB[7].tALM.tS.x3;
       "DB_M256A_Scada".tAlm.tS.tS2.x13 := "M256_Manag_IDB".M256A_IDB[7].tALM.tS.x4;
       "DB_M256A_Scada".tAlm.tS.tS2.x14 := "M256_Manag_IDB".M256A_IDB[7].tALM.tS.x5;
       "DB_M256A_Scada".tAlm.tS.tS2.x15 := "M256_Manag_IDB".M256A_IDB[7].tALM.tS.x6;
       "DB_M256A_Scada".tAlm.tS.tS2.x16 := "M256_Manag_IDB".M256A_IDB[7].tALM.tS.x7;
       "DB_M256A_Scada".tAlm.tS.tS2.x17 := "M256_Manag_IDB".M256A_IDB[7].tALM.tS.x8;
END_FUNCTION

// folder: Communication

FUNCTION "CM_Management" : Void   // FC14, LAD
{ S7_Optimized_Access := 'TRUE' }
VERSION : 0.1
   VAR_TEMP
      TMP_dDummy : DInt;
   END_VAR
   VAR_TEMP   // added for the SCL form of the ladder/FBD networks
      _w1 : Bool;
   END_VAR
BEGIN

REGION Network 1: COSTANTS
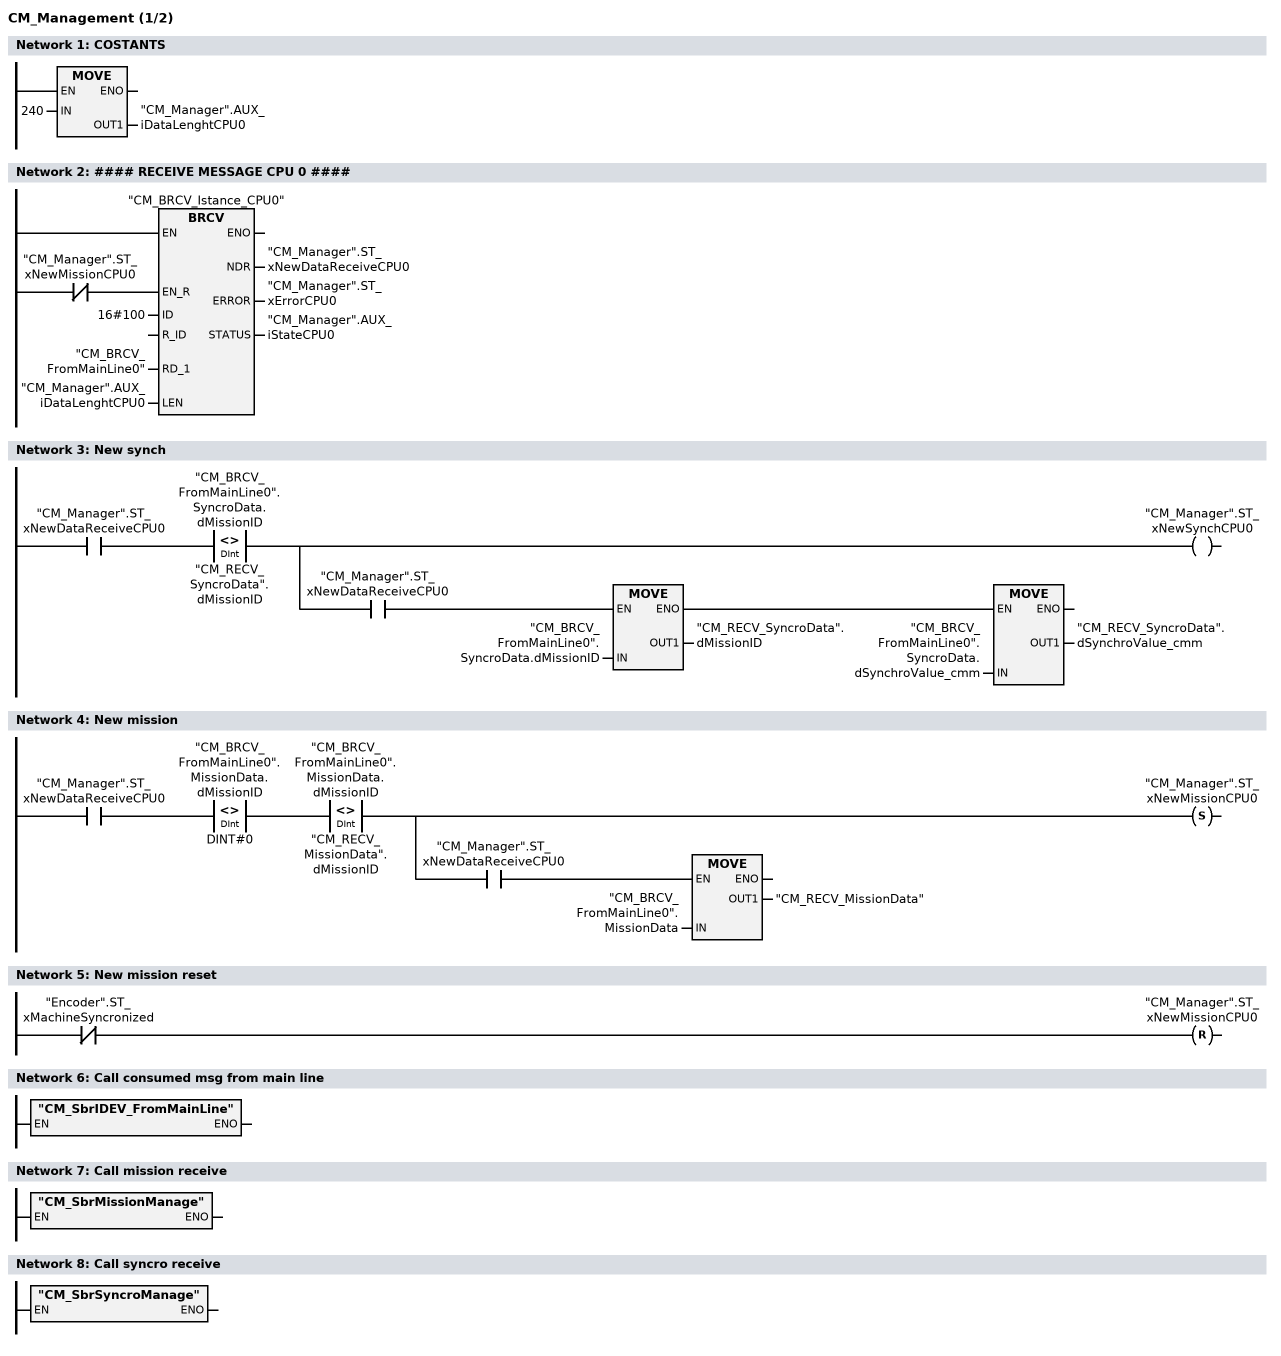
   RUNG wire#powerrail
      Move(in := 240, out1 => "CM_Manager".AUX_iDataLenghtCPU0)
   END_RUNG
   // the same network as SCL:
   "CM_Manager".AUX_iDataLenghtCPU0 := 240;
END_REGION

REGION Network 2: #### RECEIVE MESSAGE CPU 0 ####
   "CM_BRCV_Istance_CPU0"(EN_R := NOT "CM_Manager".ST_xNewMissionCPU0,   // BRCV
                          ID := 16#100,
                          RD_1 := "CM_BRCV_FromMainLine0",
                          LEN := "CM_Manager".AUX_iDataLenghtCPU0,
                          NDR => "CM_Manager".ST_xNewDataReceiveCPU0,
                          ERROR => "CM_Manager".ST_xErrorCPU0,
                          STATUS => "CM_Manager".AUX_iStateCPU0);
END_REGION

REGION Network 3: New synch
   RUNG wire#powerrail
      Contact( "CM_Manager".ST_xNewDataReceiveCPU0 )
      { S7_Templates := "SrcType := DInt" } NE_Contact(in1 := "CM_BRCV_FromMainLine0".SyncroData.dMissionID, in2 := "CM_RECV_SyncroData".dMissionID)
      wire#w1
      Coil( "CM_Manager".ST_xNewSynchCPU0 )
   END_RUNG
   RUNG wire#w1
      Contact( "CM_Manager".ST_xNewDataReceiveCPU0 )
      Move(in := "CM_BRCV_FromMainLine0".SyncroData.dMissionID, out1 => "CM_RECV_SyncroData".dMissionID)
      Move(in := "CM_BRCV_FromMainLine0".SyncroData.dSynchroValue_cmm, out1 => "CM_RECV_SyncroData".dSynchroValue_cmm)
   END_RUNG
   // the same network as SCL:
   "CM_Manager".ST_xNewSynchCPU0 := "CM_Manager".ST_xNewDataReceiveCPU0 AND ("CM_BRCV_FromMainLine0".SyncroData.dMissionID <> "CM_RECV_SyncroData".dMissionID);
   IF "CM_Manager".ST_xNewSynchCPU0 AND "CM_Manager".ST_xNewDataReceiveCPU0 THEN
       "CM_RECV_SyncroData".dMissionID := "CM_BRCV_FromMainLine0".SyncroData.dMissionID;
       "CM_RECV_SyncroData".dSynchroValue_cmm := "CM_BRCV_FromMainLine0".SyncroData.dSynchroValue_cmm;
   END_IF;
END_REGION

REGION Network 4: New mission
   RUNG wire#powerrail
      Contact( "CM_Manager".ST_xNewDataReceiveCPU0 )
      { S7_Templates := "SrcType := DInt" } NE_Contact(in1 := "CM_BRCV_FromMainLine0".MissionData.dMissionID, in2 := DINT#0)
      { S7_Templates := "SrcType := DInt" } NE_Contact(in1 := "CM_BRCV_FromMainLine0".MissionData.dMissionID, in2 := "CM_RECV_MissionData".dMissionID)
      wire#w1
      S_Coil( "CM_Manager".ST_xNewMissionCPU0 )
   END_RUNG
   RUNG wire#w1
      Contact( "CM_Manager".ST_xNewDataReceiveCPU0 )
      Move(in := "CM_BRCV_FromMainLine0".MissionData, out1 => "CM_RECV_MissionData")
   END_RUNG
   // the same network as SCL:
   #_w1 := "CM_Manager".ST_xNewDataReceiveCPU0 AND ("CM_BRCV_FromMainLine0".MissionData.dMissionID <> DINT#0) AND ("CM_BRCV_FromMainLine0".MissionData.dMissionID <> "CM_RECV_MissionData".dMissionID);
   IF #_w1 THEN "CM_Manager".ST_xNewMissionCPU0 := TRUE; END_IF;
   IF #_w1 AND "CM_Manager".ST_xNewDataReceiveCPU0 THEN
       "CM_RECV_MissionData" := "CM_BRCV_FromMainLine0".MissionData;
   END_IF;
END_REGION

REGION Network 5: New mission reset
   RUNG wire#powerrail
      I_Contact( "Encoder".ST_xMachineSyncronized )
      R_Coil( "CM_Manager".ST_xNewMissionCPU0 )
   END_RUNG
   // the same network as SCL:
   IF NOT "Encoder".ST_xMachineSyncronized THEN "CM_Manager".ST_xNewMissionCPU0 := FALSE; END_IF;
END_REGION

REGION Network 6: Call consumed msg from main line
   RUNG wire#powerrail
      "CM_SbrIDEV_FromMainLine"()
   END_RUNG
   // the same network as SCL:
   "CM_SbrIDEV_FromMainLine"();
END_REGION

REGION Network 7: Call mission receive
   RUNG wire#powerrail
      "CM_SbrMissionManage"()
   END_RUNG
   // the same network as SCL:
   "CM_SbrMissionManage"();
END_REGION

REGION Network 8: Call syncro receive
   RUNG wire#powerrail
      "CM_SbrSyncroManage"()
   END_RUNG
   // the same network as SCL:
   "CM_SbrSyncroManage"();
END_REGION

REGION Network 9: Call produced message to main line
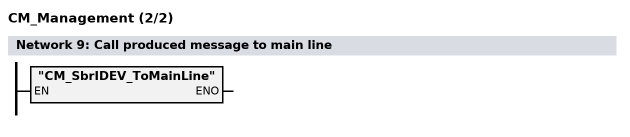
   RUNG wire#powerrail
      "CM_SbrIDEV_ToMainLine"()
   END_RUNG
   // the same network as SCL:
   "CM_SbrIDEV_ToMainLine"();
END_REGION
END_FUNCTION

FUNCTION "CM_SbrIDEV_FromMainLine" : Void   // FC15, SCL
{ S7_Optimized_Access := 'TRUE' }
VERSION : 0.1
BEGIN
   ////--------------------------------------------------------------------------------------------------------------------
   //   Copyright (c)  Bottero Spa
   //--------------------------------------------------------------
   //   Routine: ConsumedMainLine
   //       Author: Alberto Cigliutti
   //   Created: July 2016
   //--------------------------------------------------------------
   //   Description: Main line consumed message 
   //
   //   History:
   //
   ////--------------------------------------------------------------------------------------------------------------------


           "Z256".ST_xGlassBreak := "CM_IDEV_FromMainLine".xGlassBreak;
           "Z256".ST_xCycleON := "CM_IDEV_FromMainLine".xCycleON;

           IF "CM_IDEV_FromMainLine".xResetBuffers THEN
               "Z256_Manager".tInputData.xSystemReset := 1;
               "Encoder".ST_xSystemReset := 1;
           END_IF;

           IF "CM_IDEV_FromMainLine".xResetAnomaly THEN
               "Z256_hmi".tHMW.xFaultsReset := 1;
           END_IF;

    //   END_IF;
END_FUNCTION

FUNCTION "CM_SbrMissionManage" : Void   // FC16, SCL
{ S7_Optimized_Access := 'TRUE' }
VERSION : 0.1
   VAR_TEMP
      TMP_dIndex : DInt;
   END_VAR
BEGIN
   ////--------------------------------------------------------------------------------------------------------------------
   //   Copyright (c)  Bottero Spa
   //--------------------------------------------------------------
   //   Routine: CM_MissionManage
   //       Author: Alberto Cigliutti
   //   Created: July 2016
   //--------------------------------------------------------------
   //   Description: Manage the receive message
   //
   //   History:
   //
   ////--------------------------------------------------------------------------------------------------------------------

   //PLC A

   IF "CM_Manager".ST_xNewMissionCPU0 AND
       (NOT "Z256_Manager".tInputData.xNewMission) THEN


       IF (*("CM_RECV_MissionData".xPLCActive) AND*) ("Encoder".ST_xMachineSyncronized) THEN

           "Z256_Manager".tInputData.dMissionCode := "CM_RECV_MissionData".dMissionID;
           "Z256_Manager".tInputData.dMissionStart_cmm := "CM_RECV_MissionData".dMissionStart_cmm - "Encoder".AUX_dSyncroGapMainLine_cmm;
           "Z256_Manager".tInputData.dMissionEnd_cmm := "CM_RECV_MissionData".dMissionEnd_cmm - "Encoder".AUX_dSyncroGapMainLine_cmm;

           FOR #TMP_dIndex:=0 TO "CONST_dNumberOfHeadsCycle" DO
               "Z256_Manager".tInputData.rgxFireRequest[#TMP_dIndex] := "CM_RECV_MissionData".rgxFireRequest[#TMP_dIndex];
               "Z256_Manager".tInputData.rgdHeadsPosition_cmm[#TMP_dIndex] := "CM_RECV_MissionData".rgdHeadsPosition_cmm[#TMP_dIndex];
           END_FOR;

           "Z256_Manager".tInputData.xNewMission := 1;
       END_IF;

   END_IF;
END_FUNCTION

FUNCTION "CM_SbrIDEV_ToMainLine" : Void   // FC17, SCL
{ S7_Optimized_Access := 'TRUE' }
VERSION : 0.1
   VAR_TEMP
      TMP_dIndex : DInt;
   END_VAR
BEGIN
   ////--------------------------------------------------------------------------------------------------------------------
   //   Copyright (c)  Bottero Spa
   //--------------------------------------------------------------
   //   Routine: ProducedMainLine          
   //       Author: Alberto Cigliutti
   //   Created: July 2016
   //--------------------------------------------------------------
   //   Description:
   //
   //   History:
   //
   ////--------------------------------------------------------------------------------------------------------------------

   //Send request information to main line

   //Glass break in progress
   "CM_IDEV_ToMainLine".rgxStatus[0] := "CM_IDEV_FromMainLine".xGlassBreak AND (NOT "Z256_hmi".tHMW.xCutOnBreakEnabled);

   //Heads up button engaged
   "CM_IDEV_ToMainLine".rgxStatus[1] := "M256_Manag_IDB".M256A_IDB[0].INPUT_xHeadsUpIstan;

   //Bridge enabled
   "CM_IDEV_ToMainLine".rgxStatus[2] := TRUE;
   IF "M256_Manag_IDB".M256A_ST_xAllHeadStoppingFaults OR "M256_Manag_IDB".M256F_ST_xAllHeadStoppingFaults OR "M256_Manag_IDB".M256M_ST_xAllHeadStoppingFaults
       (*OR "Z256_HMI".tHMR.dProdModeActual<>3*) THEN
       "CM_IDEV_ToMainLine".rgxStatus[2] := FALSE;
   END_IF;

   //Bridge locked
   "CM_IDEV_ToMainLine".rgxStatus[3] := FALSE;

   //Cut offset calibration request (NOT USED ON MAIN LINE)
   "CM_IDEV_ToMainLine".rgxStatus[8] := FALSE;

   FOR #TMP_dIndex := 0 TO "CONST_dNumberOfHeadsCycle" DO
       "CM_IDEV_ToMainLine".rgdHeadsPositions_cmm[#TMP_dIndex] := "M256_Manag_IDB".M256M_IDB[#TMP_dIndex].AUX_dHeadActualPosition_cmm;
       "CM_IDEV_ToMainLine".rgxHeadStatus[#TMP_dIndex] := "M256_Manag_IDB".M256M_ST_xAllHeadReferred AND "Z256".INPUT_rgxHeadsInProduction[#TMP_dIndex]
       AND "Z256_hmi".tHMR.dProdModeActual=3;
       "CM_IDEV_ToMainLine".rgdHeadsPressure[#TMP_dIndex] := "M256_Manag_IDB".M256F_IDB[#TMP_dIndex].tHMW.dHeadPressure_mN;
       "CM_IDEV_ToMainLine".rgrHeadsSpace[#TMP_dIndex] := "M256_Manag_IDB".M256F_IDB[#TMP_dIndex].tHMR.rHeadUsage_km;

   END_FOR;

   //stop firing OB to have consistent data
   "CM_Manager".ST_MutingFiringOB := 1;
   FOR #TMP_dIndex := 0 TO "CONST_dNumberOfHeadsCycle" DO
       "CM_Manager".AUX_rgdHeadMissionIDInProg_Copy[#TMP_dIndex] := "M256_Manag_IDB".M256F_IDB[#TMP_dIndex].AUX_dHeadMissionIDinProg;
       "CM_Manager".AUX_rgxHeadFiringMissionInProg_Copy[#TMP_dIndex] := "M256_Manag_IDB".M256F_IDB[#TMP_dIndex].AUX_xHeadFiringMissionInProgress;
   END_FOR;
   "CM_Manager".ST_MutingFiringOB := 0;

   FOR #TMP_dIndex := 0 TO "CONST_dNumberOfHeadsCycle" DO
       "CM_IDEV_ToMainLine".dProcessingIDPlate := "CM_Manager".AUX_rgdHeadMissionIDInProg_Copy[0];
       "CM_IDEV_ToMainLine".rgxCuttingStatus[#TMP_dIndex] := "M256_Manag_IDB".M256F_IDB[#TMP_dIndex].OUTPUT_xFireON;
   END_FOR;

   //All head fire offset (NOT USED ON MAIN LINE)
   "CM_IDEV_ToMainLine".iFireOffset_OFF := 0;
   "CM_IDEV_ToMainLine".iFireOffset_ON := 0;
END_FUNCTION

FUNCTION "CM_SbrSyncroManage" : Void   // FC19, SCL
{ S7_Optimized_Access := 'TRUE' }
VERSION : 0.1
BEGIN
   ////--------------------------------------------------------------------------------------------------------------------
   //   Copyright (c)  Bottero Spa
   //--------------------------------------------------------------
   //   Routine: Syncro Manage
   //       Author: Alberto Cigliutti
   //   Created: July 2016
   //--------------------------------------------------------------
   //   Description:
   //
   //   History:
   //
   ////--------------------------------------------------------------------------------------------------------------------
   //COPY THE DATA

   //Check data received from PLC A
   IF "CM_Manager".ST_xNewSynchCPU0
       AND (NOT "Encoder".AUX_xNewSyncroReceived) THEN

       //Data valid, if PLC is active read the value 
    //   IF "CM_RECV_SyncroData".xPLCActive THEN

           "Encoder".AUX_dNewSyncroValue_cmm := "CM_RECV_SyncroData".dSynchroValue_cmm;
           "Encoder".AUX_xNewSyncroReceived := 1;

    //   END_IF;

   END_IF;
END_FUNCTION

// folder: ILx2_Blocks

FUNCTION_BLOCK "ILx2T_Control"   // FB1, SCL
{ S7_Optimized_Access := 'TRUE' }
VERSION : 1.5
   VAR_INPUT
      i_xDriveEnable : Bool;   // Enable motor current
      i_xQuickStop : Bool;   // QuickStop
      i_xHALT : Bool;   // HALT
      i_xContinue : Bool;   // Continue after HALT
      i_xFaultReset : Bool;   // Clear Error
   END_VAR
   VAR_OUTPUT
      q_byDriveState : Byte;   // Drive state
      q_xReadyToSwitchOn : Bool;   // Drive is ready to switch on (State 4)
      q_xSwitchedOn : Bool;   // Power stage is enabled (state 6 or 7)
      q_xFault : Bool;   // fault is active
      q_xWarning : Bool;   // warning is active
      q_xHALT_active : Bool;   // HALT is active
      q_xRef_OK : Bool;   // reference OK
      q_xQuickStop_Active : Bool;   // Quick Stop is active
      q_xStandstill : Bool;   // STANDSTILL
      q_xPositiveDirection : Bool;   // positive direction
      q_xNegativeDirection : Bool;   // negative direction
      q_xTargetVelocityZero : Bool;   // target velocity is zero
      q_xAccelerating : Bool;   // accelerating phase
      q_xDecelerating : Bool;   // decelerating phase
      q_xConstantVelocity : Bool;   // constant velocity
      q_woLastError : Word;   // Last Error ID (7178)
      q_woModeError : Word;   // Mode Error ID (6962)
   END_VAR
   VAR_IN_OUT
      ILx2T_Ref : "ILx2T_Ref";   // Axis reference structure
   END_VAR
   VAR
      iState : Int;   // internal state for reading error ID
      iErrorState : Int;
      inAccessID : Int;   // own access ID
      diDelayCounter : DInt;
      dwPatameterchannelError : DWord;
      WR_RetVal : Int;
      RD_RetVal : Int;
      TON_TimeOut : TON_TIME;
      xQuickStopHelper : Bool;   // Helper FAULT RESET after QuickStop
   END_VAR
   VAR_TEMP
      dwDummy : DWord;
   END_VAR
BEGIN
   // *******************************************************************************
   // Init after Restart
   // *******************************************************************************
   // Check for PLC restart (1st call of this FB)
   IF #inAccessID = 0 THEN
       #ILx2T_Ref.InitAccessID := #ILx2T_Ref.InitAccessID + 1;
       #inAccessID := #ILx2T_Ref.InitAccessID;
   END_IF;
   //******************************************************************************************************
   // Data copy into AxisRef structure
   //******************************************************************************************************
   // Processdata
   #ILx2T_Ref.i_woDriveStatus := (#ILx2T_Ref.arInputData[0] * 16#100) + #ILx2T_Ref.arInputData[1];
   #ILx2T_Ref.i_by_ModeStatus := #ILx2T_Ref.arInputData[2];
   #ILx2T_Ref.i_by_driveInput := #ILx2T_Ref.arInputData[3];
   #ILx2T_Ref.i_wo_ActionWord := (#ILx2T_Ref.arInputData[4] * 16#100) + #ILx2T_Ref.arInputData[5];
   #ILx2T_Ref.i_wo_SpecialFunctions := (#ILx2T_Ref.arInputData[6] * 16#100) + #ILx2T_Ref.arInputData[7];
   //******************************************************************************************************
   // Drive Status
   #ILx2T_Ref.stDriveStatus.HaltActive := #ILx2T_Ref.i_woDriveStatus.%X8;
   #ILx2T_Ref.stDriveStatus.reserved_Bit9 := #ILx2T_Ref.i_woDriveStatus.%X9;
   #ILx2T_Ref.stDriveStatus.reserved_Bit10 := #ILx2T_Ref.i_woDriveStatus.%X10;
   #ILx2T_Ref.stDriveStatus.reserved_Bit11 := #ILx2T_Ref.i_woDriveStatus.%X11;
   #ILx2T_Ref.stDriveStatus.reserved_Bit12 := #ILx2T_Ref.i_woDriveStatus.%X12;
   #ILx2T_Ref.stDriveStatus.x_Add := #ILx2T_Ref.i_woDriveStatus.%X13;
   #ILx2T_Ref.stDriveStatus.x_End := #ILx2T_Ref.i_woDriveStatus.%X14;
   #ILx2T_Ref.stDriveStatus.x_Err := #ILx2T_Ref.i_woDriveStatus.%X15;

   #ILx2T_Ref.stDriveStatus.state_Bit0 := #ILx2T_Ref.i_woDriveStatus.%X0;
   #ILx2T_Ref.stDriveStatus.state_Bit1 := #ILx2T_Ref.i_woDriveStatus.%X1;
   #ILx2T_Ref.stDriveStatus.state_Bit2 := #ILx2T_Ref.i_woDriveStatus.%X2;
   #ILx2T_Ref.stDriveStatus.state_Bit3 := #ILx2T_Ref.i_woDriveStatus.%X3;
   #ILx2T_Ref.stDriveStatus.reseverd_Bit4 :=#ILx2T_Ref.i_woDriveStatus.%X4;
   #ILx2T_Ref.stDriveStatus.reserved_Bit5 := #ILx2T_Ref.i_woDriveStatus.%X5;
   #ILx2T_Ref.stDriveStatus.FaultActive := #ILx2T_Ref.i_woDriveStatus.%X6;
   #ILx2T_Ref.stDriveStatus.WarningActive := #ILx2T_Ref.i_woDriveStatus.%X7;